
ScreenModuleEditorView "HMI_M_Uni_DA_mini" 1024x768
   Button "Button_2" at 95,160 size 41x40; TextOff 'Text'; PictureList "Start_M"
      on Click: InvertBit("Motor.Start_M")
      Visibility <- "Visu.view_circle"
      ObjectEnable <- "Motor.Hand"
      ProcessValue <- "Motor.Start_M"
   Circle "Circle_7" at 140,113 size 87x87
      Visibility <- "Motor.Sim"
   GraphicIOField "Graphic I/O field_1" at 146,118 size 75x75; PictureList "Pump_Down"
      Visibility <- "Type"
      ProcessValue <- "Motor.Status"
   GraphicView "Graphic view_11" at 116,89 size 30x30; Picture "service"
      Visibility <- "Motor.Trace_lock"
   GraphicIOField "Graphic I/O field_2" at 146,118 size 75x75; PictureList "Pump_Up"
      Visibility <- "Type"
      ProcessValue <- "Motor.Status"
   GraphicIOField "Graphic I/O field_3" at 146,118 size 75x75; PictureList "Pump_Left"
      Visibility <- "Type"
      ProcessValue <- "Motor.Status"
   GraphicIOField "Graphic I/O field_4" at 146,118 size 75x75; PictureList "Pump_Right"
      Visibility <- "Type"
      ProcessValue <- "Motor.Status"
   IOField "I/O field_1" at 156,190 size 55x30; FormatPattern 999.9
      Visibility <- "Motor.Analog"
      ObjectEnable <- "Motor.Hand"
      Appearance <- "Motor.Hand"
      ProcessValue <- "Motor.SP_M"
   GraphicView "Graphic view_8" at 204,176 size 30x30; Picture "force"
      Visibility <- "Motor.Force"
   GraphicView "Graphic view_12" at 134,175 size 30x30; Picture "local"
      Visibility <- "Motor.Local"
   GraphicView "Graphic view_4" at 227,128 size 38x37; Picture "z2_2"
      Visibility <- "Visu.view_circle"
   Button "Button_5" at 222,125 size 43x44; TextOff 'Text'
      on Click: ResetBit("Motor.Hand"); ResetBit("Visu.view_settings"); ResetBit("Visu.view_alm"); ResetBit("Visu.view_circle")
      Visibility <- "Visu.view_circle"
      ObjectEnable <- "Visu.view_circle"
   GraphicView "Graphic view_6" at 98,125 size 38x37; Picture "z2_1"
      Visibility <- "Visu.view_circle"
   Button "Button_6" at 95,119 size 39x44; TextOff 'Text'
      on Click: SetBit("Motor.Hand"); ResetBit("Visu.view_settings"); ResetBit("Visu.view_alm"); ResetBit("Visu.view_circle")
      Visibility <- "Visu.view_circle"
      ObjectEnable <- "Visu.view_circle"
   GraphicIOField "Graphic I/O field_5" at 146,118 size 75x75; PictureList "V_Down"
      Visibility <- "Type"
      ProcessValue <- "Motor.Status"
   GraphicIOField "Graphic I/O field_6" at 146,118 size 75x75; PictureList "V_Up"
      Visibility <- "Type"
      ProcessValue <- "Motor.Status"
   GraphicIOField "Graphic I/O field_7" at 146,118 size 75x75; PictureList "V_Left"
      Visibility <- "Type"
      ProcessValue <- "Motor.Status"
   GraphicIOField "Graphic I/O field_8" at 146,118 size 75x75; PictureList "V_Right"
      Visibility <- "Type"
      ProcessValue <- "Motor.Status"
   GraphicIOField "Graphic I/O field_9" at 146,118 size 75x75; PictureList "Z_Hor"
      Visibility <- "Type"
      ProcessValue <- "Motor.Status"
   GraphicIOField "Graphic I/O field_10" at 146,118 size 75x75; PictureList "Z_Vert"
      Visibility <- "Type"
      ProcessValue <- "Motor.Status"
   GraphicView "Graphic view_10" at 164,134 size 40x40; Picture "lock_32x32"
      Visibility <- "Motor.Lock"
   Button "Button_13" at 139,113 size 88x92; TextOff 'Text'
      on Click: InvertBit("Visu.view_circle"); ResetBit("Visu.view_alm"); ResetBit("Visu.view_settings")
   IOField "I/O field_3" at 156,91 size 55x30; FormatPattern 999.9
      Visibility <- "Motor.Analog"
      ProcessValue <- "Motor.FB_SP"
   TextField "Text field_13" at 140,72 size 85x26; Text 'Text'
      Visibility <- "Visu.view_circle"
   TextField "Text field_1" at 140,72 size 85x26; Text 'Text'
      Visibility <- "All"
   GraphicView "Graphic view_7" at 216,104 size 30x30; Picture "z2_1"
      Visibility <- "Motor.Hand"
*)

(* ===== HMI "HMI_RT_1" =====
system functions are stored by id; their names below are inferred from use

text list "Number": 1 'P1'; 2 'P2'; 3 'P3'; 4 'P11-A'; 5 'P12-A'; 6 'P13-A'; 7 'P14-I'; 8 'P15'; 9 'P4'; 10 'P6-A'; 11 'P7-A'; 12 'P21-A'; 13 'P22-A'; 14 'P10'; 15 'P11'; 16 'P12'; 17 'IE-P-02'; 18 'P26-I'; 19 'P27'; 20 'S27'; 21 'P24'; 22 'P25-A'; 23 'P25'; 24 'P29-A'; 25 'P31-A'; 26 'P33'; 27 'P25'; 28 'P26'; 29 'DP11'; 30 'DP12'; 31 'DP23'; 32 'DP65'

text list "Mode": 0 'Автомат'; 1 'Ручной'; 2 'Force'; 3 'Симуляция'; 4 'Удалённый'; 5 'Локальный'; 6 'Заблокирован'; 7 ''; 8 ''; 9 'Отключён'; 10 'Сервисный'

text list "Status": 0 'Выкл'; 1 'Вкл'; 2 'Остановка'; 3 'Запуск'; 4 'Авария ВЫКЛ'; 5 'Авария ВКЛ'; 6 'Авария QF'; 7 'Отключён'

text list "Hand": 0 'Авто'; 1 'Ручной'

text list "настройки": 0 'Настройки >>'; 1 'Настройки <<'

graphic list "Pump_Down": 1 'pump_ok'; 2 'pump_wait'; 3 'pump_wait_1'; 7 'down_stop'; 0 'pump_off'; 4 'pump'; 8 'down_start'; 9 'down_alm'

graphic list "Pump_Up": 1 'up_on'; 2 'up_wait'; 3 'up_wait'; 7 'up_stop'; 0 'up_off'; 4 'up_no'; 8 'up_start'; 9 'up_alm'

graphic list "Pump_Left": 1 'left_on'; 2 'left_wait'; 3 'left_wait_1'; 7 'left_stop'; 0 'left_off'; 4 'left_no'; 8 'left_start'; 9 'left_alm'

graphic list "Pump_Right": 1 'right_on'; 2 'right_wait'; 3 'right_wait_1'; 7 'right_stop'; 0 'right_off'; 4 'right_no'; 8 'right_start'; 9 'right_alm'

graphic list "V_Right": 1 'right_open_3x'; 2 'right_closing_3x'; 3 'right_opening_3x'; 7 'right_cl_alm_3xя'; 0 'right_close_3x'; 4 'right_no_3x'; 8 'right_op_alm_3x'; 9..100 'right_alm_3x'

graphic list "Z_Hor": 1 'h_open'; 2 'd_closing'; 3 'd_open'; 0 'v_close'; 4 'v_no'; 7..100 'down_alm_3x'

graphic list "Z_Vert": 1 'v_open'; 2 'd_closing_1'; 3 'd_opening'; 0 'h_close'; 4 'h_no'; 7..100 'h_alarm'

graphic list "V_Down": 1 'down_open_3x'; 2 'down_closing_3x'; 3 'down_opening_3x'; 7 'down_cl_alm_3xя'; 0 'down_close_3x'; 4 'down_no_3x'; 8 'down_op_alm_3x'; 9..100 'down_alm_3x'

graphic list "V_Up": 1 'up_open_3x'; 2 'up_closing_3x'; 3 'up_opening_3x'; 7 'up_cl_alm_3xя'; 0 'up_close_3x'; 4 'up_no_3x'; 8 'up_op_alm_3x'; 9 'up_alm_3x'

graphic list "V_Left": 1 'left_open_3x'; 2 'left_closing_3x'; 3 'left_opening_3x'; 7 'left_cl_alm_3xя'; 0 'left_close_3x'; 4 'left_no_3x'; 8 'left_op_alm_3x'; 9..100 'left_alm_3x'

ScreenModuleEditorView "HMI_M_Uni_DA" 1024x768
   Rectangle "Rectangle_3" at 452,30 size 168x194
      Visibility <- "Visu.view_settings"
   Rectangle "Rectangle_2" at 305,30 size 150x194
      Visibility <- "Visu.view_circle"
   GraphicIOField "Graphic I/O field_2" at 161,105 size 60x60; PictureList "Pump_Down"
      ProcessValue <- "M.Status"
      Visibility <- "Type"
   Button "Button_3" at 233,99 size 90x30; TextOff 'Авто'; TextList "Hand"
      on Click: InvertBit("M.Hand")
      ProcessValue <- "M.Hand"
      Appearance <- "M.Hand"
   Button "Button_4" at 277,143 size 45x30; TextOff 'Выкл'
      on Click: ResetBit("M.Start_M")
   Button "Button_7" at 329,60 size 122x20; TextOff 'Сервис'
      on Click: InvertBit("M.Trace_lock")
      Visibility <- "Visu.view_circle"
      Appearance <- "M.Trace_lock"
   Button "Button_8" at 329,87 size 122x20; TextOff 'Локально'
      on Click: InvertBit("M.Local")
      Visibility <- "Visu.view_circle"
      Appearance <- "M.Local"
   Button "Button_9" at 461,58 size 70x20; TextOff 'Force'
      on Click: InvertBit("M.Force")
      Visibility <- "Visu.view_settings"
      Appearance <- "M.Force"
   Button "Button_11" at 461,114 size 70x20; TextOff 'Sim'
      on Click: InvertBit("M.Sim")
      Visibility <- "Visu.view_settings"
      Appearance <- "M.Sim"
   IOField "I/O field_1" at 148,186 size 46x30; FormatPattern 999
      ProcessValue <- "M.SP_A"
      Visibility <- "M.Analog"
   IOField "I/O field_2" at 250,186 size 73x30; FormatPattern 999
      Visibility <- "M.Analog"
      ObjectEnable <- "M.Hand"
      ProcessValue <- "M.SP_M"
   Circle "Circle_4" at 598,55 size 18x18
      Visibility <- "Visu.view_settings"
      Appearance <- "M.FB_QF"
   Circle "Circle_5" at 598,83 size 18x18
      Visibility <- "Visu.view_settings"
      Appearance <- "M.FB_Run"
   TextField "Text field_4" at 535,55 size 37x18; Text 'Готов'
      Visibility <- "Visu.view_settings"
   TextField "Text field_5" at 535,83 size 56x18; Text 'В работе'
      Visibility <- "Visu.view_settings"
   IOField "I/O field_3" at 327,137 size 30x20; FormatPattern 99
      ProcessValue <- "M.Wait_On_SP"
      Visibility <- "Visu.view_circle"
   IOField "I/O field_4" at 389,137 size 30x20; FormatPattern 99
      ProcessValue <- "M.Wait_Off_SP"
      Visibility <- "Visu.view_circle"
   TextField "Text field_6" at 332,117 size 45x18; Text 'Вкл (с)'
      Visibility <- "Visu.view_circle"
   TextField "Text field_7" at 390,117 size 53x18; Text 'Выкл (с)'
      Visibility <- "Visu.view_circle"
   Button "Button_12" at 233,143 size 45x30; TextOff 'Вкл'
      on Click: SetBit("M.Start_M")
      Appearance <- "M.Start_M"
   TextField "Text field_13" at 147,60 size 177x26; Text 'Text'
   TextField "Text field_15" at 357,159 size 64x18; Text 'Задержка:'
      Visibility <- "Visu.view_circle"
   TextField "Text field_16" at 326,179 size 36x18; Text 'пуска'
      Visibility <- "Visu.view_circle"
   IOField "I/O field_6" at 381,177 size 30x20; FormatPattern 99
      ProcessValue <- "M.Delay_On_SP"
      Visibility <- "Visu.view_circle"
   IOField "I/O field_7" at 381,200 size 30x20; FormatPattern 99
      ProcessValue <- "M.Delay_Off_SP"
      Visibility <- "Visu.view_circle"
   TextField "Text field_17" at 324,200 size 56x18; Text 'останова'
      Visibility <- "Visu.view_circle"
   IOField "I/O field_8" at 411,177 size 30x20; FormatPattern 99
      ProcessValue <- "M.Delay_On_Now"
      Visibility <- "Visu.view_circle"
   IOField "I/O field_9" at 411,200 size 30x20; FormatPattern 99
      ProcessValue <- "M.Delay_Off_Now"
      Visibility <- "Visu.view_circle"
   IOField "I/O field_10" at 356,137 size 30x20; FormatPattern 99
      ProcessValue <- "M.Wait_On_Now"
      Visibility <- "Visu.view_circle"
   IOField "I/O field_11" at 419,137 size 30x20; FormatPattern 99
      ProcessValue <- "M.Wait_Off_Now"
      Visibility <- "Visu.view_circle"
   Button "Button_16" at 461,86 size 70x20; TextOff 'Impulse'
      on Click: InvertBit("M.Impulse")
      Visibility <- "Visu.view_settings"
      Appearance <- "M.Impulse"
   Circle "Circle_1" at 598,112 size 18x18
      Visibility <- "Visu.view_settings"
      Appearance <- "M.Pos_Ok"
   Circle "Circle_2" at 598,140 size 18x18
      Visibility <- "Visu.view_settings"
      Appearance <- "M.FB_Speed_Ok"
   TextField "Text field_1" at 535,112 size 53x18; Text 'Позиция'
      Visibility <- "Visu.view_settings"
   TextField "Text field_2" at 535,140 size 57x18; Text 'Скорость'
      Visibility <- "Visu.view_settings"
   Button "Button_1" at 461,143 size 70x20; TextOff 'Analog'
      on Click: InvertBit("M.Analog")
      Visibility <- "Visu.view_settings"
      Appearance <- "M.Analog"
   Button "Button_2" at 461,171 size 50x20; TextOff 'Servo'
      on Click: InvertBit("M.Servo")
      Visibility <- "Visu.view_settings"
      Appearance <- "M.Servo"
   Button "Button_5" at 461,200 size 70x20; TextOff 'Speed'
      on Click: InvertBit("M.Speed")
      Visibility <- "Visu.view_settings"
      Appearance <- "M.Speed"
   TextField "Text field_8" at 539,160 size 36x18; Text 'Servo'
      Visibility <- "Visu.view_settings"
   IOField "I/O field_5" at 541,179 size 35x20; FormatPattern 99
      ProcessValue <- "M.Delay_Servo_SP"
      Visibility <- "Visu.view_settings"
   IOField "I/O field_12" at 541,201 size 35x20; FormatPattern 99
      ProcessValue <- "M.Delay_Servo_Now"
      Visibility <- "Visu.view_settings"
   TextField "Text field_9" at 576,159 size 40x18; Text 'Speed'
      Visibility <- "Visu.view_settings"
   IOField "I/O field_13" at 581,179 size 35x20; FormatPattern 99
      ProcessValue <- "M.Delay_Speed_SP"
      Visibility <- "Visu.view_settings"
   IOField "I/O field_14" at 581,201 size 35x20; FormatPattern 99
      ProcessValue <- "M.Delay_Speed_Now"
      Visibility <- "Visu.view_settings"
   Button "Button_6" at 147,33 size 178x22; TextOff 'Настройки >>'; TextList "настройки"
      on Click: InvertBit("Visu.view_circle"); ResetBit("Visu.view_settings")
      ProcessValue <- "Visu.view_circle"
   Button "Button_10" at 329,33 size 123x22; TextOff 'Отладка >>'
      on Click: SetBit("Visu.view_settings")
      Visibility <- "Visu.view_circle"
   Button "Button_13" at 461,33 size 156x22; TextOff 'Закрыть'
      on Click: ResetBit("Visu.view_settings")
      Visibility <- "Visu.view_settings"
   GraphicIOField "Graphic I/O field_1" at 161,105 size 60x60; PictureList "Pump_Up"
      ProcessValue <- "M.Status"
      Visibility <- "Type"
   GraphicIOField "Graphic I/O field_3" at 161,105 size 60x60; PictureList "Pump_Left"
      ProcessValue <- "M.Status"
      Visibility <- "Type"
   GraphicIOField "Graphic I/O field_4" at 161,105 size 60x60; PictureList "Pump_Right"
      ProcessValue <- "M.Status"
      Visibility <- "Type"
   IOField "I/O field_15" at 194,186 size 46x30; FormatPattern 999
      ProcessValue <- "M.FB_SP"
      Visibility <- "M.Analog"
   IOField "I/O field_16" at 511,171 size 28x20; FormatPattern 9.9
      ProcessValue <- "M.Servo_DB"
      Visibility <- "Visu.view_settings"
   GraphicIOField "Graphic I/O field_5" at 161,105 size 60x60; PictureList "V_Down"
      Visibility <- "Type"
   GraphicIOField "Graphic I/O field_6" at 161,105 size 60x60; PictureList "V_Up"
      Visibility <- "Type"
   GraphicIOField "Graphic I/O field_7" at 161,105 size 60x60; PictureList "V_Left"
      Visibility <- "Type"
   GraphicIOField "Graphic I/O field_8" at 161,105 size 60x60; PictureList "V_Right"
      Visibility <- "Type"
   GraphicIOField "Graphic I/O field_9" at 161,105 size 60x60; PictureList "Z_Hor"
      Visibility <- "Type"
   GraphicIOField "Graphic I/O field_10" at 161,105 size 60x60; PictureList "Z_Vert"
      Visibility <- "Type"
   GraphicView "Graphic view_1" at 149,87 size 30x30; Picture "z2use_3"
      Visibility <- "M.Hand"
   GraphicView "Graphic view_8" at 207,86 size 30x30; Picture "force"
      Visibility <- "M.Force"
   GraphicView "Graphic view_10" at 143,128 size 50x54; Picture "lock_32x32"
      Visibility <- "M.Lock"
   GraphicView "Graphic view_11" at 199,146 size 30x30; Picture "service"
      Visibility <- "M.Trace_lock"
   GraphicView "Graphic view_12" at 179,86 size 30x30; Picture "local"
      Visibility <- "M.Local"
*)

(* ===== HMI "HMI_RT_2" =====
system functions are stored by id; their names below are inferred from use
connection "HMI_Connection_3": ETHERNET, SMART_S7_1200_OMS

HMI tags "Default tag table"
   "Clock_0.5Hz" : Bool = PLC "Clock_0.5Hz" AT %M0.7, 1 s
   "Mix_1_Clock" : Bool = PLC Mix_1_Clock AT %M10.0, 1 s
   "Mix_2_Clock" : Bool = PLC Mix_2_Clock AT %M10.1, 1 s
   "Mix_3_Clock" : Bool = PLC Mix_3_Clock AT %M10.2, 1 s
   "Logick_DB_Hand" : Bool = PLC Logick_DB.Hand AT %DB1.DBX0.1, 1 s
   "Logick_DB_Start" : Bool = PLC Logick_DB.Start AT %DB1.DBX0.0, 1 s
   "Any_Hand" : Bool = PLC Any_Hand AT %M5.0, 1 s
   "Reset_All" : Bool = PLC Reset_All AT %M3.1, 1 s
   "Logick_DB_T_Probe_SP_S" : Int = PLC Logick_DB.T_Probe.SP_S AT %DB1.DBW60, 1 s
   "Logick_DB_SP_Q" : Real = PLC Logick_DB.SP_Q AT %DB1.DBD2, 1 s
   "Logick_DB_Q" : Real = PLC Logick_DB.Q AT %DB1.DBD6, 1 s
   "Logick_DB_M" : Real = PLC Logick_DB.M AT %DB1.DBD14, 1 s
   "Logick_DB_SP_C" : Real = PLC Logick_DB.SP_C AT %DB1.DBD10, 1 s
   "Any_Alm" : Bool = PLC Any_Alm AT %M6.0, 1 s
   "Logick_DB_M_T" : Real = PLC Logick_DB.M_T AT %DB1.DBD18, 1 s
   "Logick_DB_T_Dos_SP" : Int = PLC Logick_DB.T_Dos.SP AT %DB1.DBW68, 1 s
   "Logick_DB_REQ_Calibration" : Bool = PLC Logick_DB.REQ_Calibration AT %DB1.DBX0.4, 1 s
   "Logick_DB_SP" : Real = PLC Logick_DB.SP AT %DB1.DBD22, 1 s
   "Logick_DB_L_Per_Dos" : Real = PLC Logick_DB.L_Per_Dos AT %DB1.DBD34, 1 s
   "Logick_DB_L_Percent" : Real = PLC Logick_DB.L_Percent AT %DB1.DBD42, 1 s
   "Logick_DB_T_M_SP_M" : Int = PLC Logick_DB.T_M.SP_M AT %DB1.DBW74, 1 s
   "Logick_DB_T_M_1_SP_M" : Int = PLC Logick_DB.T_M_1.SP_M AT %DB1.DBW84, 1 s
   "Logick_DB_T_M_2_SP_M" : Int = PLC Logick_DB.T_M_2.SP_M AT %DB1.DBW94, 1 s
   "Logick_DB_T_M_3_SP_M" : Int = PLC Logick_DB.T_M_3.SP_M AT %DB1.DBW104, 1 s
   "FlowMeter_DB_Full" : Real = PLC FlowMeter_DB.Full AT %DB2.DBD12, 1 s
   "Logick_DB_DD_Stop" : Bool = PLC Logick_DB.DD_Stop AT %DB1.DBX50.2, 1 s
   "Logick_DB_DD_REQ" : Bool = PLC Logick_DB.DD_REQ AT %DB1.DBX50.3, 1 s
   "Logick_DB_T_DD_Stop_SP_M" : Int = PLC Logick_DB.T_DD_Stop.SP_M AT %DB1.DBW134, 1 s
   "Logick_DB_LL_Stop" : Bool = PLC Logick_DB.LL_Stop AT %DB1.DBX50.5, 1 s
   "Logick_DB_HH_Stop" : Bool = PLC Logick_DB.HH_Stop AT %DB1.DBX50.6, 1 s
   "Logick_DB_Level_REQ" : Bool = PLC Logick_DB.Level_REQ AT %DB1.DBX50.7, 1 s
   "Logick_DB_T_Level_Stop_SP_M" : Int = PLC Logick_DB.T_Level_Stop.SP_M AT %DB1.DBW144, 1 s
   "CONFIG_Config_Use_DL" : Bool = PLC CONFIG.Config.Use_DL AT %DB10.DBX0.1, 1 s
   "CONFIG_Config_Use_DD" : Bool = PLC CONFIG.Config.Use_DD AT %DB10.DBX0.0, 1 s
   "CONFIG_Config_Use_Mix_1" : Bool = PLC CONFIG.Config.Use_Mix_1 AT %DB10.DBX0.2, 1 s
   "CONFIG_Config_Use_Mix_2" : Bool = PLC CONFIG.Config.Use_Mix_2 AT %DB10.DBX0.3, 1 s
   "CONFIG_Config_Use_Mix_3" : Bool = PLC CONFIG.Config.Use_Mix_3 AT %DB10.DBX0.4, 1 s
   "DIx_DB_M2_FB_Ready_Inverse" : Bool = PLC DIx_DB.M2_FB_Ready.Inverse AT %DB200.DBX44.3, 1 s
   "DIx_DB_DD_FB_Ready_Inverse" : Bool = PLC DIx_DB.DD_FB_Ready.Inverse AT %DB200.DBX124.3, 1 s
   "Motors_DB_DD_CMD_Sim" : Bool = PLC Motors_DB.DD.CMD.Sim AT %DB204.DBX139.2, 1 s
   "Motors_DB_Vibro_CMD_Sim" : Bool = PLC Motors_DB.Vibro.CMD.Sim AT %DB204.DBX227.2, 1 s
   "Motors_DB_DL_CMD_Sim" : Bool = PLC Motors_DB.DL.CMD.Sim AT %DB204.DBX183.2, 1 s
   "Motors_DB_Mix_1_CMD_Sim" : Bool = PLC Motors_DB.Mix_1.CMD.Sim AT %DB204.DBX7.2, 1 s
   "Motors_DB_Mix_2_CMD_Sim" : Bool = PLC Motors_DB.Mix_2.CMD.Sim AT %DB204.DBX51.2, 1 s
   "Motors_DB_Mix_3_CMD_Sim" : Bool = PLC Motors_DB.Mix_3.CMD.Sim AT %DB204.DBX95.2, 1 s
   "Motors_DB_DD_Status" : Int = PLC Motors_DB.DD.Status AT %DB204.DBW142, 1 s
   "Logick_DB_Alarm" : Word = PLC Logick_DB.Alarm AT %DB1.DBW56, 1 s
   "Motors_DB_Vibro_Status" : Int = PLC Motors_DB.Vibro.Status AT %DB204.DBW230, 1 s
   "Motors_DB_Vibro_Res_h" : DInt = PLC Motors_DB.Vibro.Res_h AT %DB204.DBD256, 1 s
   "Motors_DB_DD_Res_h" : DInt = PLC Motors_DB.DD.Res_h AT %DB204.DBD168, 1 s
   "Any_DB_Level_M" : Int = PLC Any_DB.Level_M AT %DB3.DBW0, 1 s
   "Logick_DB_Level_CMD" : Bool = PLC Logick_DB.Level_CMD AT %DB1.DBX51.0, 1 s
   "Any_DB_Flow_M" : Int = PLC Any_DB.Flow_M AT %DB3.DBW4, 1 s
   "Logick_DB_DD_CMD" : Bool = PLC Logick_DB.DD_CMD AT %DB1.DBX50.4, 1 s
   "Any_DB_DD_View" : Bool = PLC Any_DB.DD_View AT %DB3.DBX8.0, 1 s
   "Any_DB_Level_View" : Bool = PLC Any_DB.Level_View AT %DB3.DBX8.1, 1 s
   "AIx_DB_Level_Alarms_LL" : Bool = PLC AIx_DB.Level.Alarms.LL AT %DB202.DBX276.5, 1 s
   "AIx_DB_Level_Alarms_HH" : Bool = PLC AIx_DB.Level.Alarms.HH AT %DB202.DBX276.2, 1 s

HMI tags "HMI"
   "settings" : Int, internal

HMI tags "xDI"
   "DIx_DB_Vibro_FB_Ready_Signal" : Bool = PLC DIx_DB.Vibro_FB_Ready.Signal AT %DB200.DBX182.0, 1 s
   "DIx_DB_Transporter_Signal" : Bool = PLC DIx_DB.Transporter.Signal AT %DB200.DBX202.0, 1 s
   "DIx_DB_M3_FB_Run_Signal" : Bool = PLC DIx_DB.M3_FB_Run.Signal AT %DB200.DBX102.0, 1 s
   "DIx_DB_M3_FB_Ready_Signal" : Bool = PLC DIx_DB.M3_FB_Ready.Signal AT %DB200.DBX82.0, 1 s
   "DIx_DB_M2_FB_Run_Signal" : Bool = PLC DIx_DB.M2_FB_Run.Signal AT %DB200.DBX62.0, 1 s
   "DIx_DB_M2_FB_Ready_Signal" : Bool = PLC DIx_DB.M2_FB_Ready.Signal AT %DB200.DBX42.0, 1 s
   "DIx_DB_M1_FB_Run_Signal" : Bool = PLC DIx_DB.M1_FB_Run.Signal AT %DB200.DBX22.0, 1 s
   "DIx_DB_M1_FB_Ready_Signal" : Bool = PLC DIx_DB.M1_FB_Ready.Signal AT %DB200.DBX2.0, 1 s
   "DIx_DB_Dry_Run_Signal" : Bool = PLC DIx_DB.Dry_Run.Signal AT %DB200.DBX242.0, 1 s
   "DIx_DB_Dos_FB_Run_Signal" : Bool = PLC DIx_DB.Dos_FB_Run.Signal AT %DB200.DBX142.0, 1 s
   "DIx_DB_DL_FB_Ready_Signal" : Bool = PLC DIx_DB.DL_FB_Ready.Signal AT %DB200.DBX222.0, 1 s
   "DIx_DB_DD_LLS_Signal" : Bool = PLC DIx_DB.DD_LLS.Signal AT %DB200.DBX162.0, 1 s
   "DIx_DB_DD_FB_Ready_Signal" : Bool = PLC DIx_DB.DD_FB_Ready.Signal AT %DB200.DBX122.0, 1 s
   "DIx_DB_AllBlock_Signal" : Bool = PLC DIx_DB.AllBlock.Signal AT %DB200.DBX262.0, 1 s
   "DIx_DB_M1_FB_Ready_Input" : Bool = PLC DIx_DB.M1_FB_Ready.Input AT %DB200.DBX0.0, 1 s
   "DIx_DB_M1_FB_Ready_Hand" : Bool = PLC DIx_DB.M1_FB_Ready.Hand AT %DB200.DBX4.0, 1 s
   "DIx_DB_M1_FB_Ready_Start_M" : Bool = PLC DIx_DB.M1_FB_Ready.Start_M AT %DB200.DBX4.1, 1 s
   "DIx_DB_M1_FB_Ready_Inverse" : Bool = PLC DIx_DB.M1_FB_Ready.Inverse AT %DB200.DBX4.3, 1 s
   "DIx_DB_M1_FB_Ready_Filter_On_SP" : Int = PLC DIx_DB.M1_FB_Ready.Filter_On.SP AT %DB200.DBW6, 1 s
   "DIx_DB_M1_FB_Ready_Filter_Off_SP" : Int = PLC DIx_DB.M1_FB_Ready.Filter_Off.SP AT %DB200.DBW12, 1 s
   "DIx_DB_M1_FB_Run_Input" : Bool = PLC DIx_DB.M1_FB_Run.Input AT %DB200.DBX20.0, 1 s
   "DIx_DB_M1_FB_Run_Hand" : Bool = PLC DIx_DB.M1_FB_Run.Hand AT %DB200.DBX24.0, 1 s
   "DIx_DB_M1_FB_Run_Start_M" : Bool = PLC DIx_DB.M1_FB_Run.Start_M AT %DB200.DBX24.1, 1 s
   "DIx_DB_M1_FB_Run_Inverse" : Bool = PLC DIx_DB.M1_FB_Run.Inverse AT %DB200.DBX24.3, 1 s
   "DIx_DB_M1_FB_Run_Filter_On_SP" : Int = PLC DIx_DB.M1_FB_Run.Filter_On.SP AT %DB200.DBW26, 1 s
   "DIx_DB_M1_FB_Run_Filter_Off_SP" : Int = PLC DIx_DB.M1_FB_Run.Filter_Off.SP AT %DB200.DBW32, 1 s
   "DIx_DB_M2_FB_Ready_Filter_Off_SP" : Int = PLC DIx_DB.M2_FB_Ready.Filter_Off.SP AT %DB200.DBW52, 1 s
   "DIx_DB_M2_FB_Ready_Filter_On_SP" : Int = PLC DIx_DB.M2_FB_Ready.Filter_On.SP AT %DB200.DBW46, 1 s
   "DIx_DB_M2_FB_Ready_Hand" : Bool = PLC DIx_DB.M2_FB_Ready.Hand AT %DB200.DBX44.0, 1 s
   "DIx_DB_M2_FB_Ready_Start_M" : Bool = PLC DIx_DB.M2_FB_Ready.Start_M AT %DB200.DBX44.1, 1 s
   "DIx_DB_M2_FB_Ready_Input" : Bool = PLC DIx_DB.M2_FB_Ready.Input AT %DB200.DBX40.0, 1 s
   "DIx_DB_M2_FB_Run_Input" : Bool = PLC DIx_DB.M2_FB_Run.Input AT %DB200.DBX60.0, 1 s
   "DIx_DB_M2_FB_Run_Hand" : Bool = PLC DIx_DB.M2_FB_Run.Hand AT %DB200.DBX64.0, 1 s
   "DIx_DB_M2_FB_Run_Start_M" : Bool = PLC DIx_DB.M2_FB_Run.Start_M AT %DB200.DBX64.1, 1 s
   "DIx_DB_M2_FB_Run_Inverse" : Bool = PLC DIx_DB.M2_FB_Run.Inverse AT %DB200.DBX64.3, 1 s
   "DIx_DB_M2_FB_Run_Filter_On_SP" : Int = PLC DIx_DB.M2_FB_Run.Filter_On.SP AT %DB200.DBW66, 1 s
   "DIx_DB_M2_FB_Run_Filter_Off_SP" : Int = PLC DIx_DB.M2_FB_Run.Filter_Off.SP AT %DB200.DBW72, 1 s
   "DIx_DB_M3_FB_Ready_Input" : Bool = PLC DIx_DB.M3_FB_Ready.Input AT %DB200.DBX80.0, 1 s
   "DIx_DB_M3_FB_Ready_Hand" : Bool = PLC DIx_DB.M3_FB_Ready.Hand AT %DB200.DBX84.0, 1 s
   "DIx_DB_M3_FB_Ready_Start_M" : Bool = PLC DIx_DB.M3_FB_Ready.Start_M AT %DB200.DBX84.1, 1 s
   "DIx_DB_M3_FB_Ready_Inverse" : Bool = PLC DIx_DB.M3_FB_Ready.Inverse AT %DB200.DBX84.3, 1 s
   "DIx_DB_M3_FB_Ready_Filter_On_SP" : Int = PLC DIx_DB.M3_FB_Ready.Filter_On.SP AT %DB200.DBW86, 1 s
   "DIx_DB_M3_FB_Ready_Filter_Off_SP" : Int = PLC DIx_DB.M3_FB_Ready.Filter_Off.SP AT %DB200.DBW92, 1 s
   "DIx_DB_M3_FB_Run_Input" : Bool = PLC DIx_DB.M3_FB_Run.Input AT %DB200.DBX100.0, 1 s
   "DIx_DB_M3_FB_Run_Hand" : Bool = PLC DIx_DB.M3_FB_Run.Hand AT %DB200.DBX104.0, 1 s
   "DIx_DB_M3_FB_Run_Start_M" : Bool = PLC DIx_DB.M3_FB_Run.Start_M AT %DB200.DBX104.1, 1 s
   "DIx_DB_M3_FB_Run_Inverse" : Bool = PLC DIx_DB.M3_FB_Run.Inverse AT %DB200.DBX104.3, 1 s
   "DIx_DB_M3_FB_Run_Filter_On_SP" : Int = PLC DIx_DB.M3_FB_Run.Filter_On.SP AT %DB200.DBW106, 1 s
   "DIx_DB_M3_FB_Run_Filter_Off_SP" : Int = PLC DIx_DB.M3_FB_Run.Filter_Off.SP AT %DB200.DBW112, 1 s
   "DIx_DB_DD_FB_Ready_Input" : Bool = PLC DIx_DB.DD_FB_Ready.Input AT %DB200.DBX120.0, 1 s
   "DIx_DB_DD_FB_Ready_Hand" : Bool = PLC DIx_DB.DD_FB_Ready.Hand AT %DB200.DBX124.0, 1 s
   "DIx_DB_DD_FB_Ready_Start_M" : Bool = PLC DIx_DB.DD_FB_Ready.Start_M AT %DB200.DBX124.1, 1 s
   "DIx_DB_DD_FB_Ready_Filter_On_SP" : Int = PLC DIx_DB.DD_FB_Ready.Filter_On.SP AT %DB200.DBW126, 1 s
   "DIx_DB_DD_FB_Ready_Filter_Off_SP" : Int = PLC DIx_DB.DD_FB_Ready.Filter_Off.SP AT %DB200.DBW132, 1 s
   "DIx_DB_Dos_FB_Run_Input" : Bool = PLC DIx_DB.Dos_FB_Run.Input AT %DB200.DBX140.0, 1 s
   "DIx_DB_Dos_FB_Run_Hand" : Bool = PLC DIx_DB.Dos_FB_Run.Hand AT %DB200.DBX144.0, 1 s
   "DIx_DB_Dos_FB_Run_Start_M" : Bool = PLC DIx_DB.Dos_FB_Run.Start_M AT %DB200.DBX144.1, 1 s
   "DIx_DB_Dos_FB_Run_Inverse" : Bool = PLC DIx_DB.Dos_FB_Run.Inverse AT %DB200.DBX144.3, 1 s
   "DIx_DB_Dos_FB_Run_Filter_On_SP" : Int = PLC DIx_DB.Dos_FB_Run.Filter_On.SP AT %DB200.DBW146, 1 s
   "DIx_DB_Dos_FB_Run_Filter_Off_SP" : Int = PLC DIx_DB.Dos_FB_Run.Filter_Off.SP AT %DB200.DBW152, 1 s
   "DIx_DB_DD_LLS_Input" : Bool = PLC DIx_DB.DD_LLS.Input AT %DB200.DBX160.0, 1 s
   "DIx_DB_DD_LLS_Hand" : Bool = PLC DIx_DB.DD_LLS.Hand AT %DB200.DBX164.0, 1 s
   "DIx_DB_DD_LLS_Start_M" : Bool = PLC DIx_DB.DD_LLS.Start_M AT %DB200.DBX164.1, 1 s
   "DIx_DB_DD_LLS_Inverse" : Bool = PLC DIx_DB.DD_LLS.Inverse AT %DB200.DBX164.3, 1 s
   "DIx_DB_DD_LLS_Filter_On_SP" : Int = PLC DIx_DB.DD_LLS.Filter_On.SP AT %DB200.DBW166, 1 s
   "DIx_DB_DD_LLS_Filter_Off_SP" : Int = PLC DIx_DB.DD_LLS.Filter_Off.SP AT %DB200.DBW172, 1 s
   "DIx_DB_Vibro_FB_Ready_Input" : Bool = PLC DIx_DB.Vibro_FB_Ready.Input AT %DB200.DBX180.0, 1 s
   "DIx_DB_Vibro_FB_Ready_Hand" : Bool = PLC DIx_DB.Vibro_FB_Ready.Hand AT %DB200.DBX184.0, 1 s
   "DIx_DB_Vibro_FB_Ready_Start_M" : Bool = PLC DIx_DB.Vibro_FB_Ready.Start_M AT %DB200.DBX184.1, 1 s
   "DIx_DB_Vibro_FB_Ready_Inverse" : Bool = PLC DIx_DB.Vibro_FB_Ready.Inverse AT %DB200.DBX184.3, 1 s
   "DIx_DB_Vibro_FB_Ready_Filter_On_SP" : Int = PLC DIx_DB.Vibro_FB_Ready.Filter_On.SP AT %DB200.DBW186, 1 s
   "DIx_DB_Vibro_FB_Ready_Filter_Off_SP" : Int = PLC DIx_DB.Vibro_FB_Ready.Filter_Off.SP AT %DB200.DBW192, 1 s
   "DIx_DB_Transporter_Input" : Bool = PLC DIx_DB.Transporter.Input AT %DB200.DBX200.0, 1 s
   "DIx_DB_Transporter_Hand" : Bool = PLC DIx_DB.Transporter.Hand AT %DB200.DBX204.0, 1 s
   "DIx_DB_Transporter_Start_M" : Bool = PLC DIx_DB.Transporter.Start_M AT %DB200.DBX204.1, 1 s
   "DIx_DB_Transporter_Inverse" : Bool = PLC DIx_DB.Transporter.Inverse AT %DB200.DBX204.3, 1 s
   "DIx_DB_Transporter_Filter_On_SP" : Int = PLC DIx_DB.Transporter.Filter_On.SP AT %DB200.DBW206, 1 s
   "DIx_DB_Transporter_Filter_Off_SP" : Int = PLC DIx_DB.Transporter.Filter_Off.SP AT %DB200.DBW212, 1 s
   "DIx_DB_DL_FB_Ready_Input" : Bool = PLC DIx_DB.DL_FB_Ready.Input AT %DB200.DBX220.0, 1 s
   "DIx_DB_DL_FB_Ready_Hand" : Bool = PLC DIx_DB.DL_FB_Ready.Hand AT %DB200.DBX224.0, 1 s
   "DIx_DB_DL_FB_Ready_Start_M" : Bool = PLC DIx_DB.DL_FB_Ready.Start_M AT %DB200.DBX224.1, 1 s
   "DIx_DB_DL_FB_Ready_Inverse" : Bool = PLC DIx_DB.DL_FB_Ready.Inverse AT %DB200.DBX224.3, 1 s
   "DIx_DB_DL_FB_Ready_Filter_On_SP" : Int = PLC DIx_DB.DL_FB_Ready.Filter_On.SP AT %DB200.DBW226, 1 s
   "DIx_DB_DL_FB_Ready_Filter_Off_SP" : Int = PLC DIx_DB.DL_FB_Ready.Filter_Off.SP AT %DB200.DBW232, 1 s
   "DIx_DB_Dry_Run_Input" : Bool = PLC DIx_DB.Dry_Run.Input AT %DB200.DBX240.0, 1 s
   "DIx_DB_Dry_Run_Hand" : Bool = PLC DIx_DB.Dry_Run.Hand AT %DB200.DBX244.0, 1 s
   "DIx_DB_Dry_Run_Start_M" : Bool = PLC DIx_DB.Dry_Run.Start_M AT %DB200.DBX244.1, 1 s
   "DIx_DB_Dry_Run_Inverse" : Bool = PLC DIx_DB.Dry_Run.Inverse AT %DB200.DBX244.3, 1 s
   "DIx_DB_Dry_Run_Filter_On_SP" : Int = PLC DIx_DB.Dry_Run.Filter_On.SP AT %DB200.DBW246, 1 s
   "DIx_DB_Dry_Run_Filter_Off_SP" : Int = PLC DIx_DB.Dry_Run.Filter_Off.SP AT %DB200.DBW252, 1 s
   "DIx_DB_AllBlock_Filter_Off_SP" : Int = PLC DIx_DB.AllBlock.Filter_Off.SP AT %DB200.DBW272, 1 s
   "DIx_DB_AllBlock_Filter_On_SP" : Int = PLC DIx_DB.AllBlock.Filter_On.SP AT %DB200.DBW266, 1 s
   "DIx_DB_AllBlock_Inverse" : Bool = PLC DIx_DB.AllBlock.Inverse AT %DB200.DBX264.3, 1 s
   "DIx_DB_AllBlock_Start_M" : Bool = PLC DIx_DB.AllBlock.Start_M AT %DB200.DBX264.1, 1 s
   "DIx_DB_AllBlock_Hand" : Bool = PLC DIx_DB.AllBlock.Hand AT %DB200.DBX264.0, 1 s
   "DIx_DB_AllBlock_Input" : Bool = PLC DIx_DB.AllBlock.Input AT %DB200.DBX260.0, 1 s

HMI tags "xDO"
   "DOx_DB_Vibro_CMD_Q" : Bool = PLC DOx_DB.Vibro_CMD.Q AT %DB201.DBX40.2, 1 s
   "DOx_DB_M3_CMD_Q" : Bool = PLC DOx_DB.M3_CMD.Q AT %DB201.DBX20.2, 1 s
   "DOx_DB_M2_CMD_Q" : Bool = PLC DOx_DB.M2_CMD.Q AT %DB201.DBX10.2, 1 s
   "DOx_DB_M1_CMD_Q" : Bool = PLC DOx_DB.M1_CMD.Q AT %DB201.DBX0.2, 1 s
   "DOx_DB_LED_Empty_Q" : Bool = PLC DOx_DB.LED_Empty.Q AT %DB201.DBX90.2, 1 s
   "DOx_DB_LED_Dry_Run_Q" : Bool = PLC DOx_DB.LED_Dry_Run.Q AT %DB201.DBX70.2, 1 s
   "DOx_DB_LED_Alarm_Q" : Bool = PLC DOx_DB.LED_Alarm.Q AT %DB201.DBX80.2, 1 s
   "DOx_DB_KC1_CMD_Q" : Bool = PLC DOx_DB.KC1_CMD.Q AT %DB201.DBX60.2, 1 s
   "DOx_DB_DL_CMD_Q" : Bool = PLC DOx_DB.DL_CMD.Q AT %DB201.DBX50.2, 1 s
   "DOx_DB_DD_CMD_Q" : Bool = PLC DOx_DB.DD_CMD.Q AT %DB201.DBX30.2, 1 s
   "DOx_DB_M1_CMD_Start_A" : Bool = PLC DOx_DB.M1_CMD.Start_A AT %DB201.DBX0.0, 1 s
   "DOx_DB_M1_CMD_Hand" : Bool = PLC DOx_DB.M1_CMD.Hand AT %DB201.DBX2.0, 1 s
   "DOx_DB_M1_CMD_Start_M" : Bool = PLC DOx_DB.M1_CMD.Start_M AT %DB201.DBX2.1, 1 s
   "DOx_DB_M1_CMD_Simulation" : Bool = PLC DOx_DB.M1_CMD.Simulation AT %DB201.DBX2.2, 1 s
   "DOx_DB_M1_CMD_Inverse" : Bool = PLC DOx_DB.M1_CMD.Inverse AT %DB201.DBX2.3, 1 s
   "DOx_DB_M2_CMD_Start_A" : Bool = PLC DOx_DB.M2_CMD.Start_A AT %DB201.DBX10.0, 1 s
   "DOx_DB_M2_CMD_Hand" : Bool = PLC DOx_DB.M2_CMD.Hand AT %DB201.DBX12.0, 1 s
   "DOx_DB_M2_CMD_Start_M" : Bool = PLC DOx_DB.M2_CMD.Start_M AT %DB201.DBX12.1, 1 s
   "DOx_DB_M2_CMD_Simulation" : Bool = PLC DOx_DB.M2_CMD.Simulation AT %DB201.DBX12.2, 1 s
   "DOx_DB_M2_CMD_Inverse" : Bool = PLC DOx_DB.M2_CMD.Inverse AT %DB201.DBX12.3, 1 s
   "DOx_DB_M3_CMD_Start_A" : Bool = PLC DOx_DB.M3_CMD.Start_A AT %DB201.DBX20.0, 1 s
   "DOx_DB_M3_CMD_Hand" : Bool = PLC DOx_DB.M3_CMD.Hand AT %DB201.DBX22.0, 1 s
   "DOx_DB_M3_CMD_Start_M" : Bool = PLC DOx_DB.M3_CMD.Start_M AT %DB201.DBX22.1, 1 s
   "DOx_DB_M3_CMD_Simulation" : Bool = PLC DOx_DB.M3_CMD.Simulation AT %DB201.DBX22.2, 1 s
   "DOx_DB_M3_CMD_Inverse" : Bool = PLC DOx_DB.M3_CMD.Inverse AT %DB201.DBX22.3, 1 s
   "DOx_DB_DD_CMD_Start_A" : Bool = PLC DOx_DB.DD_CMD.Start_A AT %DB201.DBX30.0, 1 s
   "DOx_DB_DD_CMD_Hand" : Bool = PLC DOx_DB.DD_CMD.Hand AT %DB201.DBX32.0, 1 s
   "DOx_DB_DD_CMD_Start_M" : Bool = PLC DOx_DB.DD_CMD.Start_M AT %DB201.DBX32.1, 1 s
   "DOx_DB_DD_CMD_Simulation" : Bool = PLC DOx_DB.DD_CMD.Simulation AT %DB201.DBX32.2, 1 s
   "DOx_DB_DD_CMD_Inverse" : Bool = PLC DOx_DB.DD_CMD.Inverse AT %DB201.DBX32.3, 1 s
   "DOx_DB_Vibro_CMD_Start_A" : Bool = PLC DOx_DB.Vibro_CMD.Start_A AT %DB201.DBX40.0, 1 s
   "DOx_DB_Vibro_CMD_Hand" : Bool = PLC DOx_DB.Vibro_CMD.Hand AT %DB201.DBX42.0, 1 s
   "DOx_DB_Vibro_CMD_Start_M" : Bool = PLC DOx_DB.Vibro_CMD.Start_M AT %DB201.DBX42.1, 1 s
   "DOx_DB_Vibro_CMD_Simulation" : Bool = PLC DOx_DB.Vibro_CMD.Simulation AT %DB201.DBX42.2, 1 s
   "DOx_DB_Vibro_CMD_Inverse" : Bool = PLC DOx_DB.Vibro_CMD.Inverse AT %DB201.DBX42.3, 1 s
   "DOx_DB_DL_CMD_Start_A" : Bool = PLC DOx_DB.DL_CMD.Start_A AT %DB201.DBX50.0, 1 s
   "DOx_DB_DL_CMD_Hand" : Bool = PLC DOx_DB.DL_CMD.Hand AT %DB201.DBX52.0, 1 s
   "DOx_DB_DL_CMD_Start_M" : Bool = PLC DOx_DB.DL_CMD.Start_M AT %DB201.DBX52.1, 1 s
   "DOx_DB_DL_CMD_Simulation" : Bool = PLC DOx_DB.DL_CMD.Simulation AT %DB201.DBX52.2, 1 s
   "DOx_DB_DL_CMD_Inverse" : Bool = PLC DOx_DB.DL_CMD.Inverse AT %DB201.DBX52.3, 1 s
   "DOx_DB_KC1_CMD_Start_A" : Bool = PLC DOx_DB.KC1_CMD.Start_A AT %DB201.DBX60.0, 1 s
   "DOx_DB_KC1_CMD_Hand" : Bool = PLC DOx_DB.KC1_CMD.Hand AT %DB201.DBX62.0, 1 s
   "DOx_DB_KC1_CMD_Start_M" : Bool = PLC DOx_DB.KC1_CMD.Start_M AT %DB201.DBX62.1, 1 s
   "DOx_DB_KC1_CMD_Simulation" : Bool = PLC DOx_DB.KC1_CMD.Simulation AT %DB201.DBX62.2, 1 s
   "DOx_DB_KC1_CMD_Inverse" : Bool = PLC DOx_DB.KC1_CMD.Inverse AT %DB201.DBX62.3, 1 s
   "DOx_DB_LED_Dry_Run_Start_A" : Bool = PLC DOx_DB.LED_Dry_Run.Start_A AT %DB201.DBX70.0, 1 s
   "DOx_DB_LED_Dry_Run_Hand" : Bool = PLC DOx_DB.LED_Dry_Run.Hand AT %DB201.DBX72.0, 1 s
   "DOx_DB_LED_Dry_Run_Start_M" : Bool = PLC DOx_DB.LED_Dry_Run.Start_M AT %DB201.DBX72.1, 1 s
   "DOx_DB_LED_Dry_Run_Simulation" : Bool = PLC DOx_DB.LED_Dry_Run.Simulation AT %DB201.DBX72.2, 1 s
   "DOx_DB_LED_Dry_Run_Inverse" : Bool = PLC DOx_DB.LED_Dry_Run.Inverse AT %DB201.DBX72.3, 1 s
   "DOx_DB_LED_Alarm_Start_A" : Bool = PLC DOx_DB.LED_Alarm.Start_A AT %DB201.DBX80.0, 1 s
   "DOx_DB_LED_Alarm_Hand" : Bool = PLC DOx_DB.LED_Alarm.Hand AT %DB201.DBX82.0, 1 s
   "DOx_DB_LED_Alarm_Start_M" : Bool = PLC DOx_DB.LED_Alarm.Start_M AT %DB201.DBX82.1, 1 s
   "DOx_DB_LED_Alarm_Simulation" : Bool = PLC DOx_DB.LED_Alarm.Simulation AT %DB201.DBX82.2, 1 s
   "DOx_DB_LED_Alarm_Inverse" : Bool = PLC DOx_DB.LED_Alarm.Inverse AT %DB201.DBX82.3, 1 s
   "DOx_DB_LED_Empty_Start_A" : Bool = PLC DOx_DB.LED_Empty.Start_A AT %DB201.DBX90.0, 1 s
   "DOx_DB_LED_Empty_Hand" : Bool = PLC DOx_DB.LED_Empty.Hand AT %DB201.DBX92.0, 1 s
   "DOx_DB_LED_Empty_Start_M" : Bool = PLC DOx_DB.LED_Empty.Start_M AT %DB201.DBX92.1, 1 s
   "DOx_DB_LED_Empty_Simulation" : Bool = PLC DOx_DB.LED_Empty.Simulation AT %DB201.DBX92.2, 1 s
   "DOx_DB_LED_Empty_Inverse" : Bool = PLC DOx_DB.LED_Empty.Inverse AT %DB201.DBX92.3, 1 s
